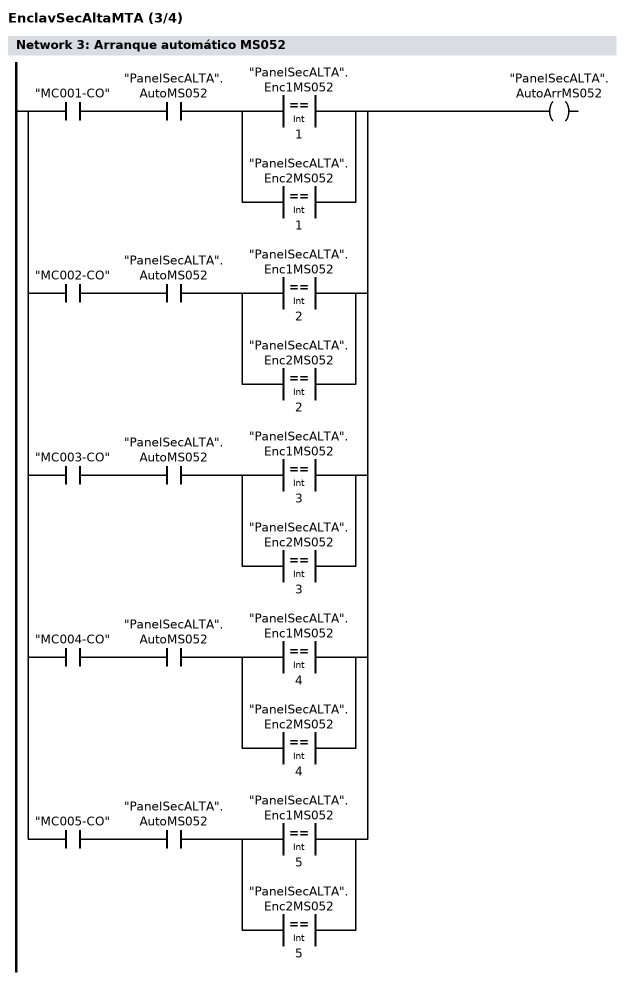
   "PanelSecALTA".AutoArrMS052 := ("MC001-CO" AND "PanelSecALTA".AutoMS052 AND (("PanelSecALTA".Enc1MS052 = 1) OR ("PanelSecALTA".Enc2MS052 = 1))) OR ("MC002-CO" AND "PanelSecALTA".AutoMS052 AND (("PanelSecALTA".Enc1MS052 = 2) OR ("PanelSecALTA".Enc2MS052 = 2))) OR ("MC003-CO" AND "PanelSecALTA".AutoMS052 AND (("PanelSecALTA".Enc1MS052 = 3) OR ("PanelSecALTA".Enc2MS052 = 3))) OR ("MC004-CO" AND "PanelSecALTA".AutoMS052 AND (("PanelSecALTA".Enc1MS052 = 4) OR ("PanelSecALTA".Enc2MS052 = 4))) OR ("MC005-CO" AND "PanelSecALTA".AutoMS052 AND (("PanelSecALTA".Enc1MS052 = 5) OR ("PanelSecALTA".Enc2MS052 = 5)));
END_REGION

REGION Network 4: Arranque automático MS053
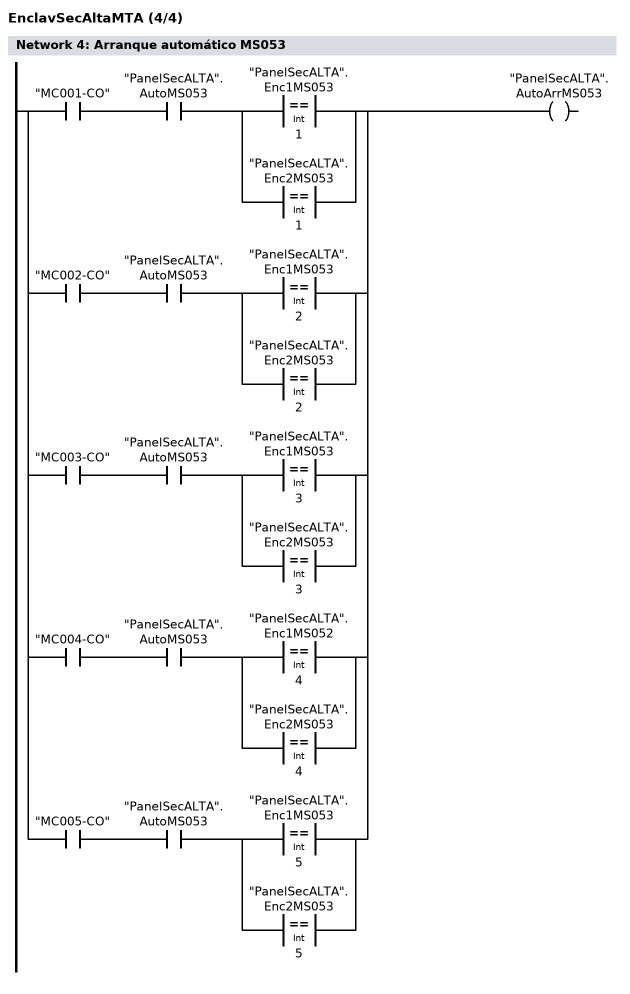
   "PanelSecALTA".AutoArrMS053 := ("MC001-CO" AND "PanelSecALTA".AutoMS053 AND (("PanelSecALTA".Enc1MS053 = 1) OR ("PanelSecALTA".Enc2MS053 = 1))) OR ("MC002-CO" AND "PanelSecALTA".AutoMS053 AND (("PanelSecALTA".Enc1MS053 = 2) OR ("PanelSecALTA".Enc2MS053 = 2))) OR ("MC003-CO" AND "PanelSecALTA".AutoMS053 AND (("PanelSecALTA".Enc1MS053 = 3) OR ("PanelSecALTA".Enc2MS053 = 3))) OR ("MC004-CO" AND "PanelSecALTA".AutoMS053 AND (("PanelSecALTA".Enc1MS052 = 4) OR ("PanelSecALTA".Enc2MS053 = 4))) OR ("MC005-CO" AND "PanelSecALTA".AutoMS053 AND (("PanelSecALTA".Enc1MS053 = 5) OR ("PanelSecALTA".Enc2MS053 = 5)));
END_REGION
END_FUNCTION

// folder: Torres de Agua/Torres Cavaleto

FUNCTION "TorresCavaletoMTA" : Void   // FC14, LAD
{ S7_Optimized_Access := 'FALSE' }
VERSION : 0.1
BEGIN

REGION Network 1: Comandos MV030 / Comandos desde Panel para MV030 - Ventilador 2 Torres de enfriamiento Cavaleto
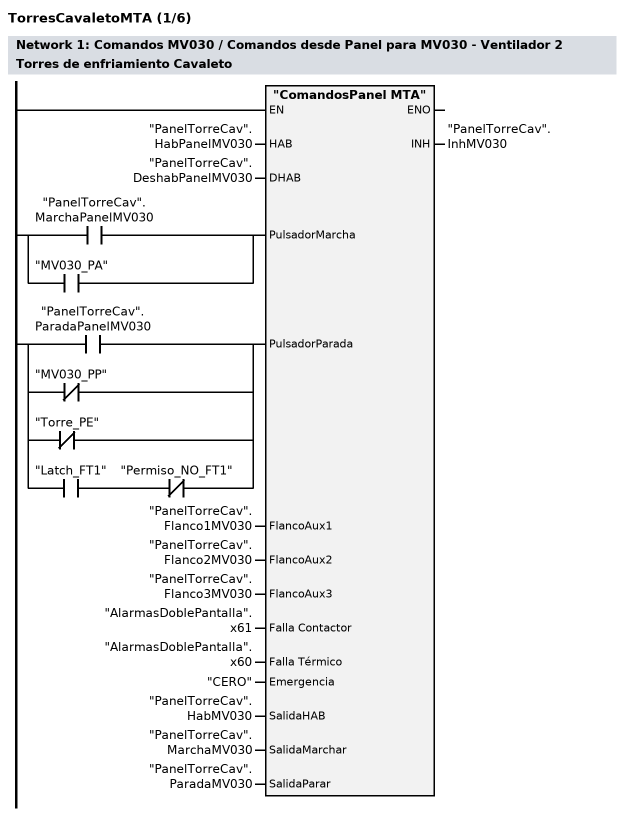
   RUNG wire#powerrail
      "ComandosPanel MTA"(PulsadorMarcha := wire#w1, PulsadorParada := wire#w2, HAB := "PanelTorreCav".HabPanelMV030, DHAB := "PanelTorreCav".DeshabPanelMV030, FlancoAux1 := "PanelTorreCav".Flanco1MV030, FlancoAux2 := "PanelTorreCav".Flanco2MV030, FlancoAux3 := "PanelTorreCav".Flanco3MV030, "Falla Contactor" := "AlarmasDoblePantalla".x61, "Falla Térmico" := "AlarmasDoblePantalla".x60, Emergencia := "CERO", SalidaHAB := "PanelTorreCav".HabMV030, SalidaMarchar := "PanelTorreCav".MarchaMV030, SalidaParar := "PanelTorreCav".ParadaMV030, INH => "PanelTorreCav".InhMV030)
   END_RUNG
   RUNG wire#powerrail
      Contact( "PanelTorreCav".MarchaPanelMV030 )
   END_RUNG wire#w1
   RUNG wire#powerrail
      Contact( "MV030_PA" )
   END_RUNG wire#w1
   RUNG wire#powerrail
      Contact( "PanelTorreCav".ParadaPanelMV030 )
   END_RUNG wire#w2
   RUNG wire#powerrail
      I_Contact( "MV030_PP" )
   END_RUNG wire#w2
   RUNG wire#powerrail
      I_Contact( "Torre_PE" )
   END_RUNG wire#w2
   RUNG wire#powerrail
      Contact( "Latch_FT1" )
      I_Contact( "Permiso_NO_FT1" )
   END_RUNG wire#w2
   // the same network as SCL:
   "ComandosPanel MTA"(HAB := "PanelTorreCav".HabPanelMV030,
                       DHAB := "PanelTorreCav".DeshabPanelMV030,
                       PulsadorMarcha := "PanelTorreCav".MarchaPanelMV030 OR "MV030_PA",
                       PulsadorParada := "PanelTorreCav".ParadaPanelMV030 OR NOT "MV030_PP" OR NOT "Torre_PE" OR ("Latch_FT1" AND NOT "Permiso_NO_FT1"),
                       FlancoAux1 := "PanelTorreCav".Flanco1MV030,
                       FlancoAux2 := "PanelTorreCav".Flanco2MV030,
                       FlancoAux3 := "PanelTorreCav".Flanco3MV030,
                       "Falla Contactor" := "AlarmasDoblePantalla".x61,
                       "Falla Térmico" := "AlarmasDoblePantalla".x60,
                       Emergencia := "CERO",
                       SalidaHAB := "PanelTorreCav".HabMV030,
                       SalidaMarchar := "PanelTorreCav".MarchaMV030,
                       SalidaParar := "PanelTorreCav".ParadaMV030,
                       INH => "PanelTorreCav".InhMV030);
END_REGION

REGION Network 2: Comandos MV031 / Comandos desde Panel para MV031 - Ventilador 1 Torres de enfriamiento Cavaleto
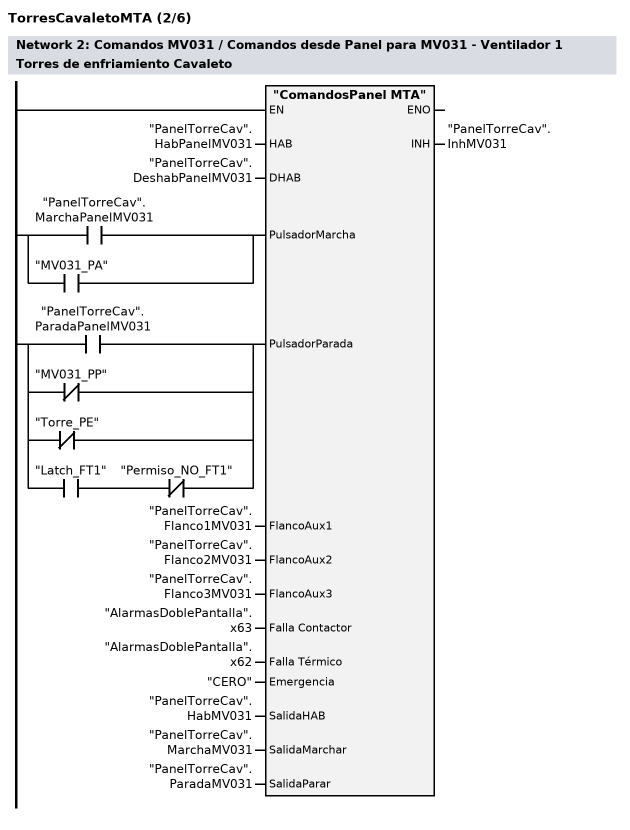
   RUNG wire#powerrail
      "ComandosPanel MTA"(PulsadorMarcha := wire#w1, PulsadorParada := wire#w2, HAB := "PanelTorreCav".HabPanelMV031, DHAB := "PanelTorreCav".DeshabPanelMV031, FlancoAux1 := "PanelTorreCav".Flanco1MV031, FlancoAux2 := "PanelTorreCav".Flanco2MV031, FlancoAux3 := "PanelTorreCav".Flanco3MV031, "Falla Contactor" := "AlarmasDoblePantalla".x63, "Falla Térmico" := "AlarmasDoblePantalla".x62, Emergencia := "CERO", SalidaHAB := "PanelTorreCav".HabMV031, SalidaMarchar := "PanelTorreCav".MarchaMV031, SalidaParar := "PanelTorreCav".ParadaMV031, INH => "PanelTorreCav".InhMV031)
   END_RUNG
   RUNG wire#powerrail
      Contact( "PanelTorreCav".MarchaPanelMV031 )
   END_RUNG wire#w1
   RUNG wire#powerrail
      Contact( "MV031_PA" )
   END_RUNG wire#w1
   RUNG wire#powerrail
      Contact( "PanelTorreCav".ParadaPanelMV031 )
   END_RUNG wire#w2
   RUNG wire#powerrail
      I_Contact( "MV031_PP" )
   END_RUNG wire#w2
   RUNG wire#powerrail
      I_Contact( "Torre_PE" )
   END_RUNG wire#w2
   RUNG wire#powerrail
      Contact( "Latch_FT1" )
      I_Contact( "Permiso_NO_FT1" )
   END_RUNG wire#w2
   // the same network as SCL:
   "ComandosPanel MTA"(HAB := "PanelTorreCav".HabPanelMV031,
                       DHAB := "PanelTorreCav".DeshabPanelMV031,
                       PulsadorMarcha := "PanelTorreCav".MarchaPanelMV031 OR "MV031_PA",
                       PulsadorParada := "PanelTorreCav".ParadaPanelMV031 OR NOT "MV031_PP" OR NOT "Torre_PE" OR ("Latch_FT1" AND NOT "Permiso_NO_FT1"),
                       FlancoAux1 := "PanelTorreCav".Flanco1MV031,
                       FlancoAux2 := "PanelTorreCav".Flanco2MV031,
                       FlancoAux3 := "PanelTorreCav".Flanco3MV031,
                       "Falla Contactor" := "AlarmasDoblePantalla".x63,
                       "Falla Térmico" := "AlarmasDoblePantalla".x62,
                       Emergencia := "CERO",
                       SalidaHAB := "PanelTorreCav".HabMV031,
                       SalidaMarchar := "PanelTorreCav".MarchaMV031,
                       SalidaParar := "PanelTorreCav".ParadaMV031,
                       INH => "PanelTorreCav".InhMV031);
END_REGION

REGION Network 3: Comandos MP014 / Comandos desde Panel para P014 - Bomba 1 Torres de enfriamiento Cavaleto
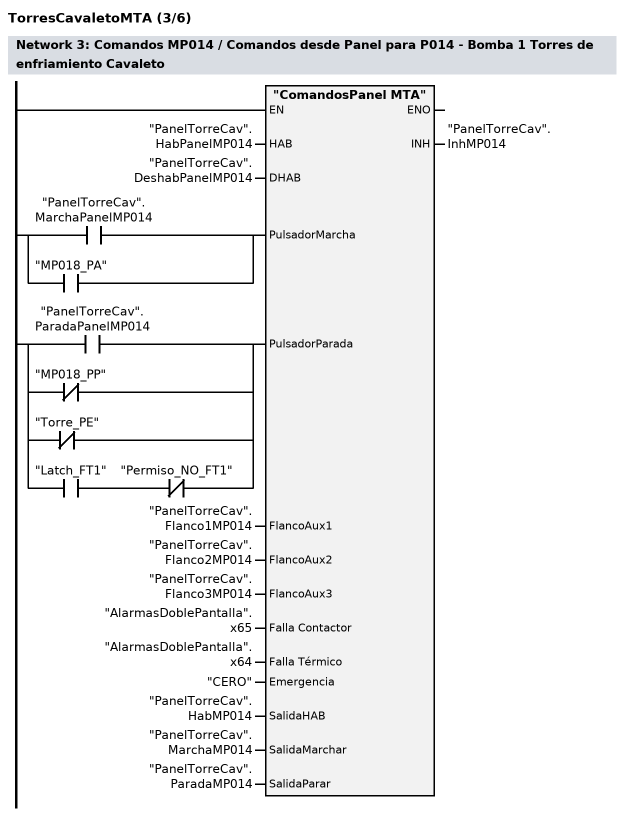
   RUNG wire#powerrail
      "ComandosPanel MTA"(PulsadorMarcha := wire#w1, PulsadorParada := wire#w2, HAB := "PanelTorreCav".HabPanelMP014, DHAB := "PanelTorreCav".DeshabPanelMP014, FlancoAux1 := "PanelTorreCav".Flanco1MP014, FlancoAux2 := "PanelTorreCav".Flanco2MP014, FlancoAux3 := "PanelTorreCav".Flanco3MP014, "Falla Contactor" := "AlarmasDoblePantalla".x65, "Falla Térmico" := "AlarmasDoblePantalla".x64, Emergencia := "CERO", SalidaHAB := "PanelTorreCav".HabMP014, SalidaMarchar := "PanelTorreCav".MarchaMP014, SalidaParar := "PanelTorreCav".ParadaMP014, INH => "PanelTorreCav".InhMP014)
   END_RUNG
   RUNG wire#powerrail
      Contact( "PanelTorreCav".MarchaPanelMP014 )
   END_RUNG wire#w1
   RUNG wire#powerrail
      Contact( "MP018_PA" )
   END_RUNG wire#w1
   RUNG wire#powerrail
      Contact( "PanelTorreCav".ParadaPanelMP014 )
   END_RUNG wire#w2
   RUNG wire#powerrail
      I_Contact( "MP018_PP" )
   END_RUNG wire#w2
   RUNG wire#powerrail
      I_Contact( "Torre_PE" )
   END_RUNG wire#w2
   RUNG wire#powerrail
      Contact( "Latch_FT1" )
      I_Contact( "Permiso_NO_FT1" )
   END_RUNG wire#w2
   // the same network as SCL:
   "ComandosPanel MTA"(HAB := "PanelTorreCav".HabPanelMP014,
                       DHAB := "PanelTorreCav".DeshabPanelMP014,
                       PulsadorMarcha := "PanelTorreCav".MarchaPanelMP014 OR "MP018_PA",
                       PulsadorParada := "PanelTorreCav".ParadaPanelMP014 OR NOT "MP018_PP" OR NOT "Torre_PE" OR ("Latch_FT1" AND NOT "Permiso_NO_FT1"),
                       FlancoAux1 := "PanelTorreCav".Flanco1MP014,
                       FlancoAux2 := "PanelTorreCav".Flanco2MP014,
                       FlancoAux3 := "PanelTorreCav".Flanco3MP014,
                       "Falla Contactor" := "AlarmasDoblePantalla".x65,
                       "Falla Térmico" := "AlarmasDoblePantalla".x64,
                       Emergencia := "CERO",
                       SalidaHAB := "PanelTorreCav".HabMP014,
                       SalidaMarchar := "PanelTorreCav".MarchaMP014,
                       SalidaParar := "PanelTorreCav".ParadaMP014,
                       INH => "PanelTorreCav".InhMP014);
END_REGION

REGION Network 4: Comandos MP015 / Comandos desde Panel para P015 - Bomba 2 Torres de enfriamiento Cavaleto
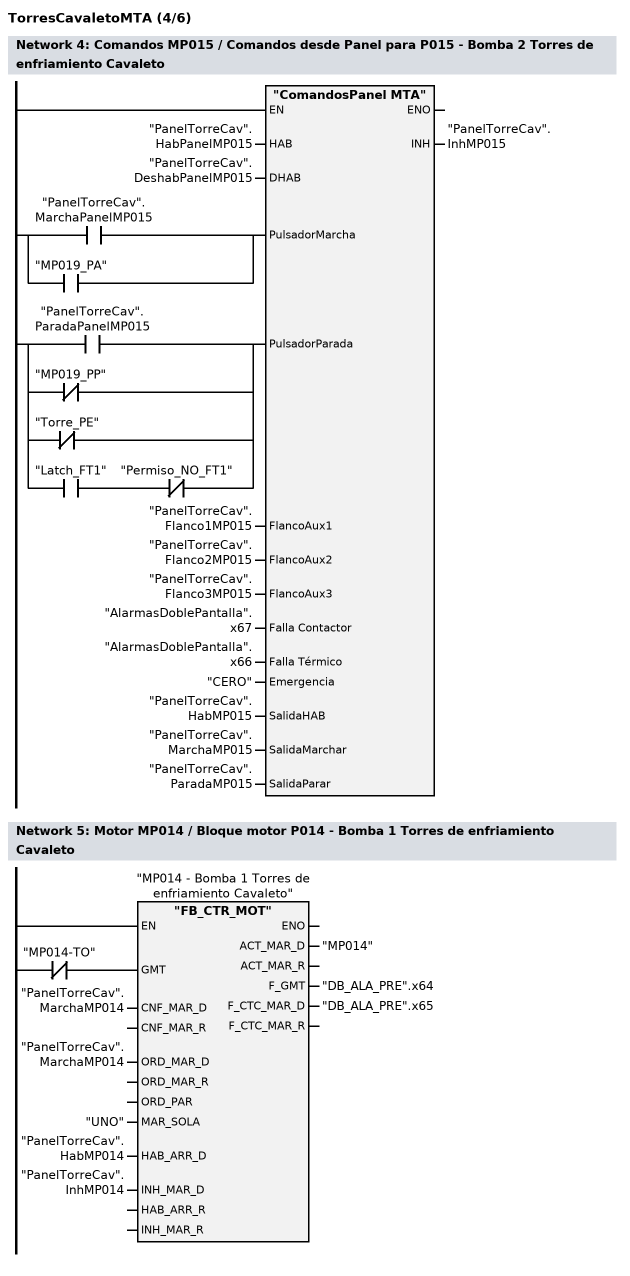
   RUNG wire#powerrail
      "ComandosPanel MTA"(PulsadorMarcha := wire#w1, PulsadorParada := wire#w2, HAB := "PanelTorreCav".HabPanelMP015, DHAB := "PanelTorreCav".DeshabPanelMP015, FlancoAux1 := "PanelTorreCav".Flanco1MP015, FlancoAux2 := "PanelTorreCav".Flanco2MP015, FlancoAux3 := "PanelTorreCav".Flanco3MP015, "Falla Contactor" := "AlarmasDoblePantalla".x67, "Falla Térmico" := "AlarmasDoblePantalla".x66, Emergencia := "CERO", SalidaHAB := "PanelTorreCav".HabMP015, SalidaMarchar := "PanelTorreCav".MarchaMP015, SalidaParar := "PanelTorreCav".ParadaMP015, INH => "PanelTorreCav".InhMP015)
   END_RUNG
   RUNG wire#powerrail
      Contact( "PanelTorreCav".MarchaPanelMP015 )
   END_RUNG wire#w1
   RUNG wire#powerrail
      Contact( "MP019_PA" )
   END_RUNG wire#w1
   RUNG wire#powerrail
      Contact( "PanelTorreCav".ParadaPanelMP015 )
   END_RUNG wire#w2
   RUNG wire#powerrail
      I_Contact( "MP019_PP" )
   END_RUNG wire#w2
   RUNG wire#powerrail
      I_Contact( "Torre_PE" )
   END_RUNG wire#w2
   RUNG wire#powerrail
      Contact( "Latch_FT1" )
      I_Contact( "Permiso_NO_FT1" )
   END_RUNG wire#w2
   // the same network as SCL:
   "ComandosPanel MTA"(HAB := "PanelTorreCav".HabPanelMP015,
                       DHAB := "PanelTorreCav".DeshabPanelMP015,
                       PulsadorMarcha := "PanelTorreCav".MarchaPanelMP015 OR "MP019_PA",
                       PulsadorParada := "PanelTorreCav".ParadaPanelMP015 OR NOT "MP019_PP" OR NOT "Torre_PE" OR ("Latch_FT1" AND NOT "Permiso_NO_FT1"),
                       FlancoAux1 := "PanelTorreCav".Flanco1MP015,
                       FlancoAux2 := "PanelTorreCav".Flanco2MP015,
                       FlancoAux3 := "PanelTorreCav".Flanco3MP015,
                       "Falla Contactor" := "AlarmasDoblePantalla".x67,
                       "Falla Térmico" := "AlarmasDoblePantalla".x66,
                       Emergencia := "CERO",
                       SalidaHAB := "PanelTorreCav".HabMP015,
                       SalidaMarchar := "PanelTorreCav".MarchaMP015,
                       SalidaParar := "PanelTorreCav".ParadaMP015,
                       INH => "PanelTorreCav".InhMP015);
END_REGION

REGION Network 5: Motor MP014 / Bloque motor P014 - Bomba 1 Torres de enfriamiento Cavaleto
   RUNG wire#powerrail
      "MP014 - Bomba 1 Torres de enfriamiento Cavaleto"(CNF_MAR_D := "PanelTorreCav".MarchaMP014, CNF_MAR_R :=, ORD_MAR_D := "PanelTorreCav".MarchaMP014, ORD_MAR_R :=, ORD_PAR :=, MAR_SOLA := "UNO", HAB_ARR_D := "PanelTorreCav".HabMP014, INH_MAR_D := "PanelTorreCav".InhMP014, HAB_ARR_R :=, INH_MAR_R :=, ACT_MAR_D => "MP014", ACT_MAR_R =>, F_GMT => "DB_ALA_PRE".x64, F_CTC_MAR_D => "DB_ALA_PRE".x65, F_CTC_MAR_R =>, GMT := wire#w1)
   END_RUNG
   RUNG wire#powerrail
      I_Contact( "MP014-TO" )
   END_RUNG wire#w1
   // the same network as SCL:
   "MP014 - Bomba 1 Torres de enfriamiento Cavaleto"(GMT := NOT "MP014-TO",   // "FB_CTR_MOT"
                           CNF_MAR_D := "PanelTorreCav".MarchaMP014,
                           ORD_MAR_D := "PanelTorreCav".MarchaMP014,
                           MAR_SOLA := "UNO",
                           HAB_ARR_D := "PanelTorreCav".HabMP014,
                           INH_MAR_D := "PanelTorreCav".InhMP014,
                           ACT_MAR_D => "MP014",
                           F_GMT => "DB_ALA_PRE".x64,
                           F_CTC_MAR_D => "DB_ALA_PRE".x65);
END_REGION

REGION Network 6: Motor MP015 / Bloque motor P015 - Bomba 2 Torres de enfriamiento Cavaleto
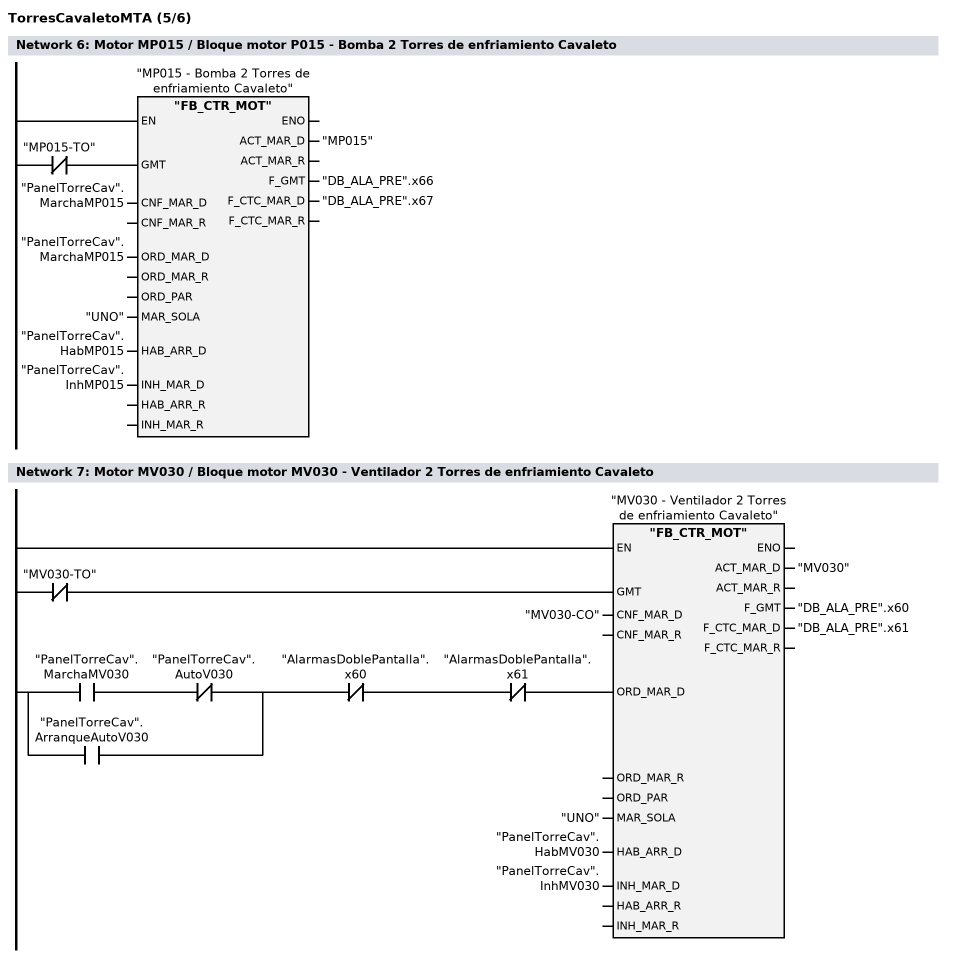
   RUNG wire#powerrail
      "MP015 - Bomba 2 Torres de enfriamiento Cavaleto"(CNF_MAR_D := "PanelTorreCav".MarchaMP015, CNF_MAR_R :=, ORD_MAR_D := "PanelTorreCav".MarchaMP015, ORD_MAR_R :=, ORD_PAR :=, MAR_SOLA := "UNO", HAB_ARR_D := "PanelTorreCav".HabMP015, INH_MAR_D := "PanelTorreCav".InhMP015, HAB_ARR_R :=, INH_MAR_R :=, ACT_MAR_D => "MP015", ACT_MAR_R =>, F_GMT => "DB_ALA_PRE".x66, F_CTC_MAR_D => "DB_ALA_PRE".x67, F_CTC_MAR_R =>, GMT := wire#w1)
   END_RUNG
   RUNG wire#powerrail
      I_Contact( "MP015-TO" )
   END_RUNG wire#w1
   // the same network as SCL:
   "MP015 - Bomba 2 Torres de enfriamiento Cavaleto"(GMT := NOT "MP015-TO",   // "FB_CTR_MOT"
                           CNF_MAR_D := "PanelTorreCav".MarchaMP015,
                           ORD_MAR_D := "PanelTorreCav".MarchaMP015,
                           MAR_SOLA := "UNO",
                           HAB_ARR_D := "PanelTorreCav".HabMP015,
                           INH_MAR_D := "PanelTorreCav".InhMP015,
                           ACT_MAR_D => "MP015",
                           F_GMT => "DB_ALA_PRE".x66,
                           F_CTC_MAR_D => "DB_ALA_PRE".x67);
END_REGION

REGION Network 7: Motor MV030 / Bloque motor MV030 - Ventilador 2 Torres de enfriamiento Cavaleto
   RUNG wire#powerrail
      "MV030 - Ventilador 2 Torres de enfriamiento Cavaleto"(GMT := wire#w1, ORD_MAR_D := wire#w3, CNF_MAR_D := "MV030-CO", CNF_MAR_R :=, ORD_MAR_R :=, ORD_PAR :=, MAR_SOLA := "UNO", HAB_ARR_D := "PanelTorreCav".HabMV030, INH_MAR_D := "PanelTorreCav".InhMV030, HAB_ARR_R :=, INH_MAR_R :=, ACT_MAR_D => "MV030", ACT_MAR_R =>, F_GMT => "DB_ALA_PRE".x60, F_CTC_MAR_D => "DB_ALA_PRE".x61, F_CTC_MAR_R =>)
   END_RUNG
   RUNG wire#powerrail
      I_Contact( "MV030-TO" )
   END_RUNG wire#w1
   RUNG wire#powerrail
      Contact( "PanelTorreCav".MarchaMV030 )
      I_Contact( "PanelTorreCav".AutoV030 )
      wire#w2
      I_Contact( "AlarmasDoblePantalla".x60 )
      I_Contact( "AlarmasDoblePantalla".x61 )
   END_RUNG wire#w3
   RUNG wire#powerrail
      Contact( "PanelTorreCav".ArranqueAutoV030 )
   END_RUNG wire#w2
   // the same network as SCL:
   "MV030 - Ventilador 2 Torres de enfriamiento Cavaleto"(GMT := NOT "MV030-TO",   // "FB_CTR_MOT"
                           CNF_MAR_D := "MV030-CO",
                           ORD_MAR_D := (("PanelTorreCav".MarchaMV030 AND NOT "PanelTorreCav".AutoV030) OR "PanelTorreCav".ArranqueAutoV030) AND NOT "AlarmasDoblePantalla".x60 AND NOT "AlarmasDoblePantalla".x61,
                           MAR_SOLA := "UNO",
                           HAB_ARR_D := "PanelTorreCav".HabMV030,
                           INH_MAR_D := "PanelTorreCav".InhMV030,
                           ACT_MAR_D => "MV030",
                           F_GMT => "DB_ALA_PRE".x60,
                           F_CTC_MAR_D => "DB_ALA_PRE".x61);
END_REGION

REGION Network 8: Motor MV031 / Bloque motorMV031 - Ventilador 1 Torres de enfriamiento Cavaleto
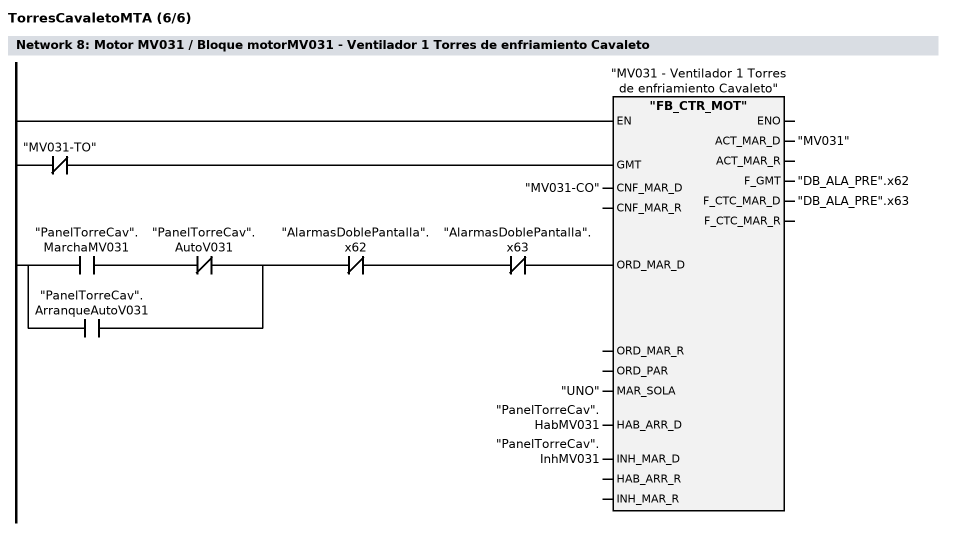
   RUNG wire#powerrail
      "MV031 - Ventilador 1 Torres de enfriamiento Cavaleto"(GMT := wire#w1, ORD_MAR_D := wire#w3, CNF_MAR_D := "MV031-CO", CNF_MAR_R :=, ORD_MAR_R :=, ORD_PAR :=, MAR_SOLA := "UNO", HAB_ARR_D := "PanelTorreCav".HabMV031, INH_MAR_D := "PanelTorreCav".InhMV031, HAB_ARR_R :=, INH_MAR_R :=, ACT_MAR_D => "MV031", ACT_MAR_R =>, F_GMT => "DB_ALA_PRE".x62, F_CTC_MAR_D => "DB_ALA_PRE".x63, F_CTC_MAR_R =>)
   END_RUNG
   RUNG wire#powerrail
      I_Contact( "MV031-TO" )
   END_RUNG wire#w1
   RUNG wire#powerrail
      Contact( "PanelTorreCav".MarchaMV031 )
      I_Contact( "PanelTorreCav".AutoV031 )
      wire#w2
      I_Contact( "AlarmasDoblePantalla".x62 )
      I_Contact( "AlarmasDoblePantalla".x63 )
   END_RUNG wire#w3
   RUNG wire#powerrail
      Contact( "PanelTorreCav".ArranqueAutoV031 )
   END_RUNG wire#w2
   // the same network as SCL:
   "MV031 - Ventilador 1 Torres de enfriamiento Cavaleto"(GMT := NOT "MV031-TO",   // "FB_CTR_MOT"
                           CNF_MAR_D := "MV031-CO",
                           ORD_MAR_D := (("PanelTorreCav".MarchaMV031 AND NOT "PanelTorreCav".AutoV031) OR "PanelTorreCav".ArranqueAutoV031) AND NOT "AlarmasDoblePantalla".x62 AND NOT "AlarmasDoblePantalla".x63,
                           MAR_SOLA := "UNO",
                           HAB_ARR_D := "PanelTorreCav".HabMV031,
                           INH_MAR_D := "PanelTorreCav".InhMV031,
                           ACT_MAR_D => "MV031",
                           F_GMT => "DB_ALA_PRE".x62,
                           F_CTC_MAR_D => "DB_ALA_PRE".x63);
END_REGION
END_FUNCTION

// folder: Torres de Agua/Torres Chillers

FUNCTION "TorresAutoMTA" : Void   // FC9, LAD
{ S7_Optimized_Access := 'FALSE' }
VERSION : 0.1
BEGIN

REGION Network 1: Lectura Temperatura de Torres Chillers
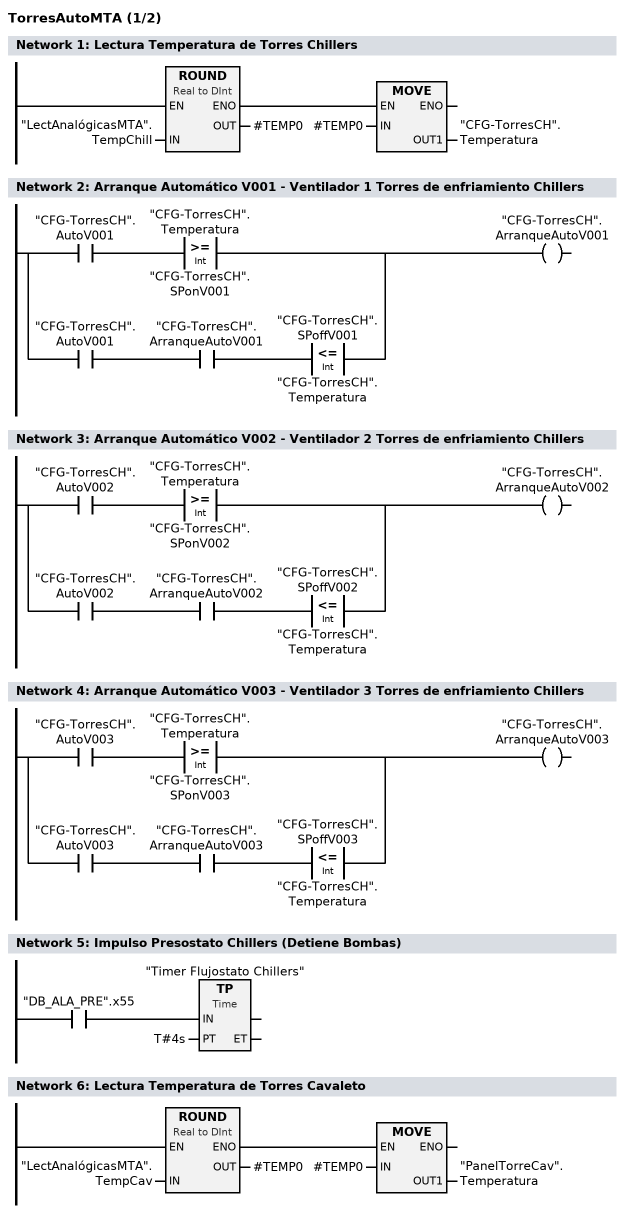
   RUNG wire#powerrail
      { S7_Templates := "[SrcType := Real, DestType := DInt]"; S7_GenerateENO := "TRUE" } Round(in := "LectAnalógicasMTA".TempChill, out => #TEMP0)
      { S7_GenerateENO := "TRUE" } Move(in := #TEMP0, out1 => "CFG-TorresCH".Temperatura)
   END_RUNG
   // the same network as SCL:
   // ENO of a box is taken as its EN; it also drops when the box reports an error
   #TEMP0 := ROUND("LectAnalógicasMTA".TempChill);
   "CFG-TorresCH".Temperatura := #TEMP0;
END_REGION

REGION Network 2: Arranque Automático V001 - Ventilador 1 Torres de enfriamiento Chillers
   "CFG-TorresCH".ArranqueAutoV001 := ("CFG-TorresCH".AutoV001 AND ("CFG-TorresCH".Temperatura >= "CFG-TorresCH".SPonV001)) OR ("CFG-TorresCH".AutoV001 AND "CFG-TorresCH".ArranqueAutoV001 AND ("CFG-TorresCH".SPoffV001 <= "CFG-TorresCH".Temperatura));
END_REGION

REGION Network 3: Arranque Automático V002 - Ventilador 2 Torres de enfriamiento Chillers
   "CFG-TorresCH".ArranqueAutoV002 := ("CFG-TorresCH".AutoV002 AND ("CFG-TorresCH".Temperatura >= "CFG-TorresCH".SPonV002)) OR ("CFG-TorresCH".AutoV002 AND "CFG-TorresCH".ArranqueAutoV002 AND ("CFG-TorresCH".SPoffV002 <= "CFG-TorresCH".Temperatura));
END_REGION

REGION Network 4: Arranque Automático V003 - Ventilador 3 Torres de enfriamiento Chillers
   "CFG-TorresCH".ArranqueAutoV003 := ("CFG-TorresCH".AutoV003 AND ("CFG-TorresCH".Temperatura >= "CFG-TorresCH".SPonV003)) OR ("CFG-TorresCH".AutoV003 AND "CFG-TorresCH".ArranqueAutoV003 AND ("CFG-TorresCH".SPoffV003 <= "CFG-TorresCH".Temperatura));
END_REGION

REGION Network 5: Impulso Presostato Chillers (Detiene Bombas)
   "Timer Flujostato Chillers".TP(in := "DB_ALA_PRE".x55, pt := T#4s);
END_REGION

REGION Network 6: Lectura Temperatura de Torres Cavaleto
   RUNG wire#powerrail
      { S7_Templates := "[SrcType := Real, DestType := DInt]"; S7_GenerateENO := "TRUE" } Round(in := "LectAnalógicasMTA".TempCav, out => #TEMP0)
      { S7_GenerateENO := "TRUE" } Move(in := #TEMP0, out1 => "PanelTorreCav".Temperatura)
   END_RUNG
   // the same network as SCL:
   // ENO of a box is taken as its EN; it also drops when the box reports an error
   #TEMP0 := ROUND("LectAnalógicasMTA".TempCav);
   "PanelTorreCav".Temperatura := #TEMP0;
END_REGION

REGION Network 7: Arranque Automático MV030 - Ventilador 1 Torres de enfriamiento Cavaleto
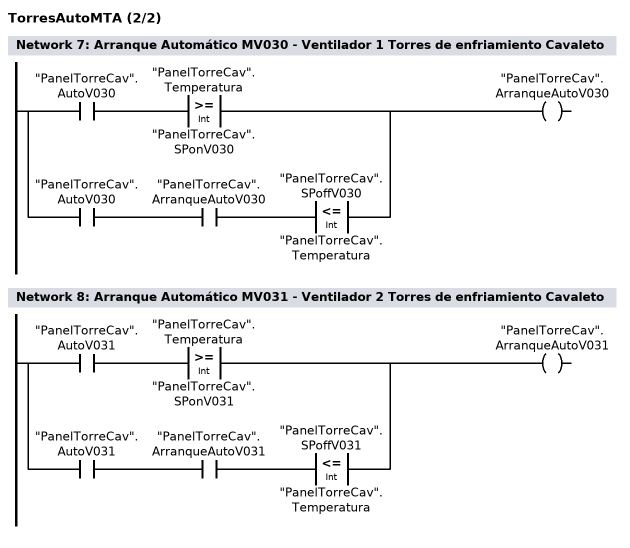
   "PanelTorreCav".ArranqueAutoV030 := ("PanelTorreCav".AutoV030 AND ("PanelTorreCav".Temperatura >= "PanelTorreCav".SPonV030)) OR ("PanelTorreCav".AutoV030 AND "PanelTorreCav".ArranqueAutoV030 AND ("PanelTorreCav".SPoffV030 <= "PanelTorreCav".Temperatura));
END_REGION

REGION Network 8: Arranque Automático MV031 - Ventilador 2 Torres de enfriamiento Cavaleto
   "PanelTorreCav".ArranqueAutoV031 := ("PanelTorreCav".AutoV031 AND ("PanelTorreCav".Temperatura >= "PanelTorreCav".SPonV031)) OR ("PanelTorreCav".AutoV031 AND "PanelTorreCav".ArranqueAutoV031 AND ("PanelTorreCav".SPoffV031 <= "PanelTorreCav".Temperatura));
END_REGION
END_FUNCTION

(* ===== HMI "HMI_RT_3" =====
connection "Conexión2-PLC_1": ETHERNET, SIMATIC S7 300/400 MPI

HMI tags "AlarmasMTA"
   "AlarmasWord0" : Int, 1 s
   "AlarmasWord1" : Int, 1 s
   "AlarmasWord2" : Int, 1 s
   "AlarmasWord3" : Int, 1 s
   "AlarmasWord4" : Int, 1 s
   "AlarmasWord5" : Int, 1 s
   "AlarmasWord6" : Int, 1 s
   "AlarmasWord7" : Int, 1 s
   "AlarmasWord8" : Int, 1 s
   "Rec0" : Int, 1 s
   "Rec1" : Int, 1 s
   "Rec2" : Int, 1 s
   "Rec3" : Int, 1 s
   "Rec4" : Int, 1 s
   "Rec5" : Int, 1 s
   "Rec6" : Int, 1 s
   "Rec7" : Int, 1 s
   "Rec8" : Int, 1 s
   "AlarmasWord9" : Int, 1 s
   "AlarmasWord10" : Int, 1 s
   "AlarmasWord11" : Int, 1 s
   "AlarmasWord12" : Int, 1 s
   "AlarmasWord13" : Int, 1 s
   "AlarmasWord14" : Int, 1 s
   "Rec9" : Int, 1 s
   "Rec10" : Int, 1 s
   "Rec11" : Int, 1 s
   "Rec12" : Int, 1 s
   "Rec13" : Int, 1 s
   "Rec14" : Int, 1 s
   "AlarmasWord1(1)" : Int, 1 s
   "AlarmasWord15" : Int, 1 s
   "Rec15" : Int, 1 s
   "EncendidoPLC" : Bool, 1 s

HMI tags "AutoTorresChillers"
   "AutoV001" : Bool, 1 s
   "AutoV002" : Bool, 1 s
   "AutoV003" : Bool, 1 s
   "SP-ON-V001" : Int, 1 s
   "SP-ON-V002" : Int, 1 s
   "SP-ON-V003" : Int, 1 s
   "SP-OFF-V001" : Int, 1 s
   "SP-OFF-V002" : Int, 1 s
   "SP-OFF-V003" : Int, 1 s
   "TemperaturatorresCH" : Real, 1 s

HMI tags "CFG-Analog-MTA"
   "PresiónALTA" : Real, 1 s
   "PresiónBAJA" : Real, 1 s
   "TempCAV" : Real, 1 s
   "TempCH" : Real, 1 s
   "CFG-ALtaHH" : Real, 1 s
   "CFG-ALtaH" : Real, 1 s
   "CFG-ALtaL" : Real, 1 s
   "CFG-ALtaLL" : Real, 1 s
   "CFG-BajaHH" : Real, 1 s
   "CFG-BajaH" : Real, 1 s
   "CFG-BajaL" : Real, 1 s
   "CFG-BajaLL" : Real, 1 s

HMI tags "ChillersMTA"
   "HabMT007" : Bool, 1 s
   "HabMT008" : Bool, 1 s
   "HabMT009" : Bool, 1 s
   "HabMT010" : Bool, 1 s
   "DesMT007" : Bool, 1 s
   "DesMT008" : Bool, 1 s
   "DesMT009" : Bool, 1 s
   "DesMT010" : Bool, 1 s
   "MarchaMT007" : Bool, 1 s
   "MarchaMT008" : Bool, 1 s
   "MarchaMT009" : Bool, 1 s
   "MarchaMT010" : Bool, 1 s
   "ParadaMT007" : Bool, 1 s
   "ParadaMT008" : Bool, 1 s
   "ParadaMT009" : Bool, 1 s
   "ParadaMT010" : Bool, 1 s
   "Habilitación-CH-SOP-GR" : Bool, 1 s
   "Habilitación-CH-SOP-CH" : Bool, 1 s
   "Habilitación-CH-ENV-GR" : Bool, 1 s
   "Habilitación-CH-ENV-CH" : Bool, 1 s
   "Alarma1-CH-SOP-GR" : Bool, 1 s
   "Alarma2-CH-SOP-GR" : Bool, 1 s
   "RUN-CH-SOP-GR" : Bool, 1 s
   "MAX-CH-SOP-GR" : Bool, 1 s
   "AnimaciónMT007" : Byte, 1 s
   "AnimaciónMT008" : Byte, 1 s
   "AnimaciónMT009" : Byte, 1 s
   "AnimaciónMT010" : Byte, 1 s
   "AnimaciónMP010" : Byte, 1 s
   "AnimaciónMP011" : Byte, 1 s
   "AnimaciónMP012" : Byte, 1 s
   "AnimaciónMP013" : Byte, 1 s
   "HabMP010" : Bool, 1 s
   "HabMP011" : Bool, 1 s
   "HabMP012" : Bool, 1 s
   "HabMP013" : Bool, 1 s
   "HabMP018" : Bool, 1 s
   "HabMP019" : Bool, 1 s
   "DesMP010" : Bool, 1 s
   "DesMP011" : Bool, 1 s
   "DesMP012" : Bool, 1 s
   "DesMP013" : Bool, 1 s
   "DesMP018" : Bool, 1 s
   "DesMP019" : Bool, 1 s
   "MarchaMP010" : Bool, 1 s
   "MarchaMP011" : Bool, 1 s
   "MarchaMP012" : Bool, 1 s
   "MarchaMP013" : Bool, 1 s
   "MarchaMP018" : Bool, 1 s
   "MarchaMP019" : Bool, 1 s
   "ParadaMP010" : Bool, 1 s
   "ParadaMP011" : Bool, 1 s
   "ParadaMP012" : Bool, 1 s
   "ParadaMP013" : Bool, 1 s
   "ParadaMP018" : Bool, 1 s
   "ParadaMP019" : Bool, 1 s
   "AnimaciónMP018" : Byte, 1 s
   "AnimaciónMP019" : Byte, 1 s
   "DesV001" : Bool, 1 s
   "DesV002" : Bool, 1 s
   "HabV001" : Bool, 1 s
   "HabV002" : Bool, 1 s
   "MarchaV001" : Bool, 1 s
   "MarchaV002" : Bool, 1 s
   "ParadaV001" : Bool, 1 s
   "ParadaV002" : Bool, 1 s
   "AnimaciónV001" : Byte, 1 s
   "AnimaciónV002" : Byte, 1 s
   "VentiladoresMTA" : Bool, internal
   "MAX-CH-ENV-GR" : Bool, 1 s
   "RUN-CH-ENV-GR" : Bool, 1 s
   "Alarma2-CH-ENV-GR" : Bool, 1 s
   "Alarma1-CH-ENV-GR" : Bool, 1 s
   "SirenaM1" : Bool, 1 s
   "SirenaM2" : Bool, 1 s
   "SirenaM3" : Bool, 1 s
   "SirenaM4" : Bool, 1 s
   "AnimaciónV003" : Byte, 1 s
   "HabV003" : Bool, 1 s
   "DesV003" : Bool, 1 s
   "MarchaV003" : Bool, 1 s
   "ParadaV003" : Bool, 1 s
   "BombaTorreON" : Bool, 1 s
   "SirenaM5" : Bool, 1 s
   "SirenaChillers" : Bool, 1 s
   "SirenaM6" : Bool, 1 s
   "SirenaM7" : Bool, 1 s
   "SirenaM8" : Bool, 1 s
   "SirenaM9" : Bool, 1 s
   "SirenaM10" : Bool, 1 s
   "AlarmaNueva" : Bool, 1 s
   "AlarmaPresente" : Bool, 1 s
   "SinAlarmas" : Bool, 1 s
   "AlarmaAceite-CH-ENV-CH" : Bool, 1 s
   "AlarmaTemp-CH-ENV-CH" : Bool, 1 s
   "RUN-CH-ENV-CH" : Bool, 1 s
   "VerCh1MTA" : Bool, internal
   "VerCh2MTA" : Bool, internal
   "VerCh3MTA" : Bool, internal
   "VerCh4MTA" : Bool, internal
   "AlarmaPRUEBA" : DWord, 1 s
   "Presosato" : Bool, 1 s
   "CH-SOP-CH-CTC1ON" : Bool, 1 s
   "CH-SOP-CH-CTC2ON" : Bool, 1 s
   "CH-SOP-CH-TERM1" : Bool, 1 s
   "CH-SOP-CH-TERM2" : Bool, 1 s
   "CH-ENV-CH-ACT" : Bool, 1 s
   "CH-ENV-CH-TEMP" : Bool, 1 s
   "CH-ENV-CH-TERM" : Bool, 1 s
   "CH-ENV-CH-RUN" : Bool, 1 s
   "BombaTorreON2" : Bool, 1 s
   "HabV001(1)" : Bool, 1 s
   "HabV002(1)" : Bool, 1 s
   "HabV003(1)" : Bool, 1 s
   "HabV4" : Bool, 1 s
   "MarchaV001(1)" : Bool, 1 s
   "MarchaV002(1)" : Bool, 1 s
   "MarchaV003(1)" : Bool, 1 s
   "ParadaV001(1)" : Bool, 1 s
   "ParadaV002(1)" : Bool, 1 s
   "ParadaV003(1)" : Bool, 1 s
   "AnimaMenuV001" : Int, 1 s
   "AnimaMenuV002" : Int, 1 s
   "AnimaMenuV003" : Int, 1 s
   "DeshV001" : Bool, 1 s
   "DeshV002" : Bool, 1 s
   "DeshV003" : Bool, 1 s